// TIA Portal project "StepTimeAnalysis" (V16) (continued)
REGION Network 25: Archive values Step 9
   "DB_HMI".ARG1_Seq1_S9 := "IDB_Arg_Seq_1_DB".Step9.X;
END_REGION

REGION Network 26: Archive values Step 10
   "DB_HMI".ARG1_Seq1_S10 := "IDB_Arg_Seq_1_DB".Step10.X;
END_REGION

REGION Network 27: Archive values Step 11
   "DB_HMI".ARG1_Seq1_S11 := "IDB_Arg_Seq_1_DB".Step11.X;
END_REGION

REGION Network 28: Archive values Step 12
   "DB_HMI".ARG1_Seq1_S12 := "IDB_Arg_Seq_1_DB".Step12.X;
END_REGION

REGION Network 29: Archive values Step 13
   "DB_HMI".ARG1_Seq1_S13 := "IDB_Arg_Seq_1_DB".Step13.X;
END_REGION

REGION Network 30: Archive values Step 14
   "DB_HMI".ARG1_Seq1_S14 := "IDB_Arg_Seq_1_DB".Step14.X;
END_REGION

REGION Network 31: Archive values Step 15
   "DB_HMI".ARG1_Seq1_S15 := "IDB_Arg_Seq_1_DB".Step15.X;
END_REGION

REGION Network 32: Archive values Step 16
   "DB_HMI".ARG1_Seq1_S16 := "IDB_Arg_Seq_1_DB".Step16.X;
END_REGION

REGION Network 33: Archive values Step 17
   "DB_HMI".ARG1_Seq1_S17 := "IDB_Arg_Seq_1_DB".Step17.X;
END_REGION

REGION Network 34: Archive values Step 18
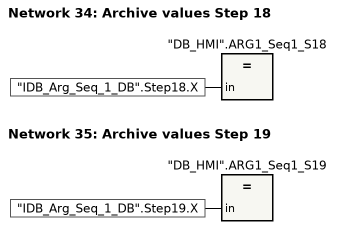
   "DB_HMI".ARG1_Seq1_S18 := "IDB_Arg_Seq_1_DB".Step18.X;
END_REGION

REGION Network 35: Archive values Step 19
   "DB_HMI".ARG1_Seq1_S19 := "IDB_Arg_Seq_1_DB".Step19.X;
END_REGION

REGION Network 36 (SCL): Set Busy
   IF
       "IDB_Arg_Seq_1_DB".Step2.X OR
       "IDB_Arg_Seq_1_DB".Step3.X OR
       "IDB_Arg_Seq_1_DB".Step4.X OR
       "IDB_Arg_Seq_1_DB".Step5.X OR
       "IDB_Arg_Seq_1_DB".Step6.X OR
       "IDB_Arg_Seq_1_DB".Step7.X OR
       "IDB_Arg_Seq_1_DB".Step8.X OR
       "IDB_Arg_Seq_1_DB".Step9.X OR
       "IDB_Arg_Seq_1_DB".Step10.X OR
       "IDB_Arg_Seq_1_DB".Step11.X OR
       "IDB_Arg_Seq_1_DB".Step12.X OR
       "IDB_Arg_Seq_1_DB".Step13.X OR
       "IDB_Arg_Seq_1_DB".Step14.X OR
       "IDB_Arg_Seq_1_DB".Step15.X OR
       "IDB_Arg_Seq_1_DB".Step16.X OR
       "IDB_Arg_Seq_1_DB".Step17.X OR
       "IDB_Arg_Seq_1_DB".Step18.X OR
       "IDB_Arg_Seq_1_DB".Step19.X THEN
       "DB_HMI".ARG1_Seq1_Status_Busy := TRUE;
   ELSIF "IDB_Arg_Seq_1_DB"."Step1: Init (Idle)".X THEN
       "DB_HMI".ARG1_Seq1_Status_Busy := FALSE;
   END_IF;
END_REGION

REGION Network 37 (SCL): When Stepper Sequence runs completely
   IF "IDB_Arg_Seq_1_DB".Trans10.TS = TRUE OR "IDB_Arg_Seq_1_DB".Trans21.TS = TRUE THEN
       "DB_Process_Var".Branch_Complete := TRUE;
       "DB_Process_Var".Car_Type_Ready := "DB_Process_Var".Car_Type_inProduction;
       "DB_Process_Var".Car_Type_inProduction := 0;
       "DB_Process_Var".Car_Type_inProduction_Text := '';
       "DB_Process_Var".Car_ReadyToShift := TRUE;
       "DB_HMI".ARG1_Seq1_inProduction := 0;
   END_IF;
   IF "IDB_Arg_Seq_1_DB".Trans1.TS = TRUE OR "IDB_Arg_Seq_1_DB".Trans11.TS = TRUE THEN
       "DB_Process_Var".Branch_Complete := FALSE;
       "DB_Process_Var".ReadyNewCar := 0;
   END_IF;
END_REGION

REGION Network 38 (SCL): Write Data in the Sending Box
   //IF "DB_Process_Var".Branch_Complete = TRUE AND "DB_PLC1_Receiving".ReceivingBox.Station_Idle = TRUE THEN
   IF "IDB_Arg_Seq_1_DB".Trans10.TS = TRUE OR "IDB_Arg_Seq_1_DB".Trans21.TS = TRUE THEN
       "DB_PLC1_Sending".SendBoxForward.Planned_PT_Red := "DB_HMI".ARG1_Seq1_Calculated_PT_Red;
       "DB_PLC1_Sending".SendBoxForward.Planned_PT_Green := "DB_HMI".ARG1_Seq1_Calculated_PT_Green;
       "DB_PLC1_Sending".SendBoxForward.Planned_PT_Blue := "DB_HMI".ARG1_Seq1_Calculated_PT_Blue;

       "DB_PLC1_Sending".SendBoxForward.Measuered_PT_Red := "DB_HMI".ARG1_Seq1_Messured_PT_Red;
       "DB_PLC1_Sending".SendBoxForward.Measuered_PT_Green := "DB_HMI".ARG1_Seq1_Messured_PT_Green;
       "DB_PLC1_Sending".SendBoxForward.Measuered_PT_Blue := "DB_HMI".ARG1_Seq1_Messured_PT_Blue;

       "DB_PLC1_Sending".SendBoxForward.Type := "DB_Process_Var".Car_Type_Ready;

       "DB_PLC1_Receiving".ReceivingBoxForward.Type := 0;
   END_IF;
END_REGION

REGION Network 39 (SCL)
   //IF "DB_Process_Var".Branch_Complete = TRUE AND "DB_PLC1_Receiving".ReceivingBox.Station_Idle = TRUE THEN
    //   "DB_Process_Var".ready_new_car := TRUE;
   //END_IF;
END_REGION

REGION Network 40 (SCL): When car is shifted
   IF "DB_Process_Var".Data_Put_Done = TRUE THEN
       "DB_Process_Var".Car_Type_Ready := 0;
       "DB_PLC1_Sending".SendBoxForward.Type := 0;
       "DB_Process_Var".Car_ReadyToShift := FALSE;
       "DB_Process_Var".ReadyNewCar := 1;

       //"DB_PLC1_Receiving".ReceivingBoxForward.Type := 0;
   END_IF;
END_REGION
END_FUNCTION

FUNCTION "FC_Com" : Void   // FC2, FBD
{ S7_Optimized_Access := 'TRUE' }
VERSION : 0.1
BEGIN

REGION Network 1: Communication PLC1 -> PLC2
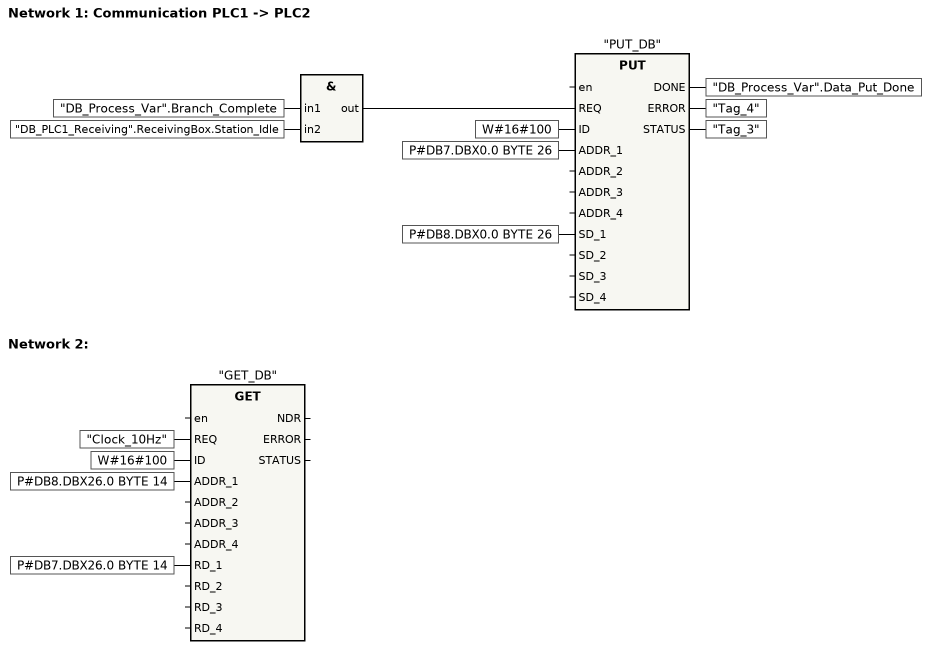
   "PUT_DB"(REQ := "DB_Process_Var".Branch_Complete AND "DB_PLC1_Receiving".ReceivingBox.Station_Idle,   // PUT
            ID := W#16#100,
            ADDR_1 := P#DB7.DBX0.0 BYTE 26,
            SD_1 := P#DB8.DBX0.0 BYTE 26,
            DONE => "DB_Process_Var".Data_Put_Done,
            ERROR => "Tag_4",
            STATUS => "Tag_3");
END_REGION

REGION Network 2
   "GET_DB"(REQ := "Clock_10Hz", ID := W#16#100, ADDR_1 := P#DB8.DBX26.0 BYTE 14, RD_1 := P#DB7.DBX26.0 BYTE 14);   // GET
END_REGION
END_FUNCTION

FUNCTION "FC_PT_Calc" : Void   // FC3, SCL
{ S7_Optimized_Access := 'TRUE' }
VERSION : 0.1
   VAR_TEMP
      i : Int;
   END_VAR
   VAR CONSTANT
      sequenceNO : Int := 9;
      Null : Time := T#0MS;
   END_VAR
BEGIN
   "DB_HMI".ARG1_Seq1_Calculated_PT_Red := #Null;
   "DB_HMI".ARG1_Seq1_Calculated_PT_Green := #Null;
   "DB_HMI".ARG1_Seq1_Calculated_PT_Blue := #Null;

   "DB_HMI".ARG1_Seq1_Messured_PT_Red := #Null;
   "DB_HMI".ARG1_Seq1_Messured_PT_Green := #Null;
   "DB_HMI".ARG1_Seq1_Messured_PT_Blue := #Null;

   FOR #i := 2 TO #sequenceNO + 1 DO
       //Calculated Production Time
       "DB_HMI".ARG1_Seq1_Calculated_PT_Red := "DB_HMI".ARG1_Seq1_Calculated_PT_Red + "DB_Profile".time_Red[#i];
       "DB_HMI".ARG1_Seq1_Calculated_PT_Green := "DB_HMI".ARG1_Seq1_Calculated_PT_Green + "DB_Profile".time_Green[#i];
       "DB_HMI".ARG1_Seq1_Calculated_PT_Blue := "DB_HMI".ARG1_Seq1_Calculated_PT_Blue + "DB_Profile".time_Blue[#i];
       //Messured Production Time
       IF "DB_Process_Var".Car_Type_inProduction = 3 THEN
           "DB_HMI".ARG1_Seq1_Messured_PT_Red := "DB_HMI".ARG1_Seq1_Messured_PT_Red + "DB_Process_Var".Step_Times[#i];
       ELSIF "DB_Process_Var".Car_Type_inProduction = 4 THEN
           "DB_HMI".ARG1_Seq1_Messured_PT_Green := "DB_HMI".ARG1_Seq1_Messured_PT_Green + "DB_Process_Var".Step_Times[#i];
       ELSIF "DB_Process_Var".Car_Type_inProduction = 6 THEN
           "DB_HMI".ARG1_Seq1_Messured_PT_Blue := "DB_HMI".ARG1_Seq1_Messured_PT_Blue + "DB_Process_Var".Step_Times[#i];
       END_IF;
   END_FOR;

   //Add Time of previous Stations
   "DB_HMI".ARG1_Seq1_Calculated_PT_Red := "DB_HMI".ARG1_Seq1_Calculated_PT_Red + "DB_PLC1_Receiving".ReceivingBoxForward.Planned_PT_Red;
   "DB_HMI".ARG1_Seq1_Calculated_PT_Green := "DB_HMI".ARG1_Seq1_Calculated_PT_Green + "DB_PLC1_Receiving".ReceivingBoxForward.Planned_PT_Green;
   "DB_HMI".ARG1_Seq1_Calculated_PT_Blue := "DB_HMI".ARG1_Seq1_Calculated_PT_Blue + "DB_PLC1_Receiving".ReceivingBoxForward.Planned_PT_Blue;

   "DB_HMI".ARG1_Seq1_Messured_PT_Red := "DB_HMI".ARG1_Seq1_Messured_PT_Red + "DB_PLC1_Receiving".ReceivingBoxForward.Measuered_PT_Red;
   "DB_HMI".ARG1_Seq1_Messured_PT_Green := "DB_HMI".ARG1_Seq1_Messured_PT_Green + "DB_PLC1_Receiving".ReceivingBoxForward.Measuered_PT_Green;
   "DB_HMI".ARG1_Seq1_Messured_PT_Blue := "DB_HMI".ARG1_Seq1_Messured_PT_Blue + "DB_PLC1_Receiving".ReceivingBoxForward.Measuered_PT_Blue;
END_FUNCTION

FUNCTION "FC_Global_Status" : Void   // FC4, SCL
{ S7_Optimized_Access := 'TRUE' }
VERSION : 0.1
   VAR_TEMP
      global_auto : Bool;
      global_man : Bool;
      test2 : Bool;
      test : Bool;
      i : Int;
   END_VAR
BEGIN
   IF "DB_Process_Var".Auto_Mode = TRUE THEN
       "DB_PLC1_Sending".SendBox.Mode_PLC1 := 1;
   ELSIF "DB_Process_Var".Man_Mode = TRUE THEN
       "DB_PLC1_Sending".SendBox.Mode_PLC1 := 2;
   ELSE
       "DB_PLC1_Sending".SendBox.Mode_PLC1 := 0;
   END_IF;

   IF "DB_Process_Var".Station_Nr = 1 THEN
       IF "DB_PLC1_Sending".SendBox.Mode_PLC1 = 1 AND "DB_PLC1_Receiving".ReceivingBox.Mode_PLC2 = 1 AND "DB_PLC1_Receiving".ReceivingBox.Mode_PLC3 = 1 AND "DB_PLC1_Receiving".ReceivingBox.Mode_PLC4 = 1 AND "DB_PLC1_Receiving".ReceivingBox.Mode_PLC5 = 1 THEN
           "DB_HMI".Global_Status_Auto := TRUE;
           "DB_HMI".Global_Status_Man := FALSE;
       ELSIF "DB_PLC1_Sending".SendBox.Mode_PLC1 = 0 AND "DB_PLC1_Receiving".ReceivingBox.Mode_PLC2 = 0 AND "DB_PLC1_Receiving".ReceivingBox.Mode_PLC3 = 0 AND "DB_PLC1_Receiving".ReceivingBox.Mode_PLC4 = 0 AND "DB_PLC1_Receiving".ReceivingBox.Mode_PLC5 = 0 THEN
           "DB_HMI".Global_Status_Auto := FALSE;
           "DB_HMI".Global_Status_Man := FALSE;
       ELSE
           "DB_HMI".Global_Status_Man := TRUE;
           "DB_HMI".Global_Status_Auto := FALSE;
       END_IF;
   END_IF;


   //Global Selection
   "DB_PLC1_Receiving".ReceivingBoxForward.Type := "DB_HMI".Global_selection;
END_FUNCTION

ORGANIZATION_BLOCK "Main"   // OB1, LAD, ProgramCycle
TITLE = "Main Program Sweep (Cycle)"
{ S7_Optimized_Access := 'TRUE' }
VERSION : 0.1
   VAR_INPUT
      Initial_Call : Bool;   // Initial call of this OB
      Remanence : Bool;   // =True, if remanent data are available
   END_VAR
   VAR_TEMP
      test : Bool;
   END_VAR
BEGIN

REGION Network 1: Call ARG_1
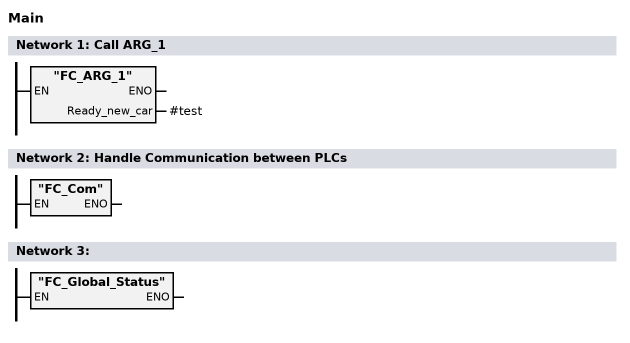
   RUNG wire#powerrail
      "FC_ARG_1"(Ready_new_car => #test)
   END_RUNG
   // the same network as SCL:
   "FC_ARG_1"(Ready_new_car => #test);
END_REGION

REGION Network 2: Handle Communication between PLCs
   RUNG wire#powerrail
      "FC_Com"()
   END_RUNG
   // the same network as SCL:
   "FC_Com"();
END_REGION

REGION Network 3
   RUNG wire#powerrail
      "FC_Global_Status"()
   END_RUNG
   // the same network as SCL:
   "FC_Global_Status"();
END_REGION
END_ORGANIZATION_BLOCK

// folder: LGF/4 Math operations

FUNCTION "LGF_RandomRange_Dint" : DInt   // FC10013, SCL
TITLE = LGF_RandomRange_DInt
{ S7_Optimized_Access := 'TRUE' }
AUTHOR : Siemens_Digital_Industries
FAMILY : LGF
NAME : LGF_RandomRange_DInt
// This function generates random numbers in defined limits (Datatype DInt)
   VAR_INPUT
      minValue : DInt;   // minimal Value random can reach / Minimum value of the range of the random number
      maxValue : DInt;   // maximal Value random can reach / Maximum value of the range of the random number
   END_VAR
   VAR_OUTPUT
      error : Bool;   // Error if true
      status : Word;   // Status of the function
      subfunctionStatus : Word;   // Status or return value of called FB's, FCs and system blocks
   END_VAR
   VAR_TEMP
      tempTime : DTL;   // System time
      tempNanoSecondInDWord : DWord;   // UDINT converted to DWORD for access to individual bytes
      tempTimeStatus : Word;   // Status of the instruction RD_SYS_T
      tempRandomValue : DWord;   // Random-start-value
      tempNormReal : Real;   // Normalized value
   END_VAR
   // Ret_Val : Returns random DInt number in a predefined range
   VAR CONSTANT
      ZERO : DInt := 0;   // Zero value in case of error
      MAX_UDINT : UDInt := 4294967295 ;   // Maximum UDINT value
      SUB_STATUS_NO_ERROR : Word := 16#0000;   // Status: sub function call ends without error
      STATUS_FINISHED_NO_ERROR : Word := 16#0000;   // Status: Execution finished without errors
      ERR_MAX_LESS_MIN : Word := 16#8200;   // Error: The maximum limit number is smaller than the minimum limit number
      ERR_RD_SYS_T : Word := 16#8600;   // Error: System function Read system time returned an error
   END_VAR
BEGIN
   REGION Block info header
     //=============================================================================
     // SIEMENS AG / (c)Copyright 2017
     //-----------------------------------------------------------------------------
     // Title:            LGF_RandomRange_DInt
     // Comment/Function: This function generates random numbers in defined limits (Datatype DInt)
     // Library/Family:   LGF(Library General Functions)
     // Author:           Siemens Digital Industry Support
     // Tested with:      S7-PLCSIM Advanced V2.0 SP1
     // Engineering:      TIA Portal V15 Update 2
     // Restrictions:     ENO disabled - error handling done by error and status
     // Requirements:     PLC (S7-1200 / S7-1500)
     //-------------------------------------------------------------------------------
     // Change log table:
     // Version  | Date       | Expert in charge       | Changes applied
     //----------|------------|------------------------|------------------------------
     // 01.00.00 19.08.2015  Siemens Industry Online Support
     //                      First released version
     // 01.00.01 02.01.2017  Siemens Industry Online Support
     //                      Upgrade: TIA Portal V14 Update 1
     // 01.00.02 17.08.2018  Siemens Industry Online Support
     //                      Upgrade: TIA V15 Update 2
     // 01.00.03 23.11.2018  Siemens Industry Online Support
     //                      Upgrade: TIA V15.1
     // 01.01.00 09.10.2019  Siemens Industry Presales Support
     //                      Renamed from "LGF_RandomInt" to "LGF_RandomRange_DInt"
     //                      change random datatype from int to dint
     //                      Regions, commens and costants are added
     // 03.00.00 23.04.2020  Siemens Industry Support
     //                      Set version to V3.0.0, harmonize the version of the whole library
     //=============================================================================
   END_REGION

   REGION Validation
     // Check if the maximal Value is less than the minimal value
     IF (#minValue > #maxValue) THEN
       #error := true;
       #status := #ERR_MAX_LESS_MIN;
       #subfunctionStatus := #SUB_STATUS_NO_ERROR;
       #LGF_RandomRange_Dint := #ZERO;
       RETURN;
     END_IF;

     // Read system time
     #tempTimeStatus := INT_TO_WORD(RD_SYS_T(#tempTime));

     // Check return variable for error
     IF (#tempTimeStatus <> #SUB_STATUS_NO_ERROR) THEN
       #error := true;
       #status := #ERR_RD_SYS_T;
       #subfunctionStatus := #tempTimeStatus;
       #LGF_RandomRange_Dint := #ZERO;
       RETURN;
     END_IF;
   END_REGION

   REGION Calculating random number
     // Converting to double word so individual bytes can be addressed
     #tempNanoSecondInDWord := UDINT_TO_DWORD(#tempTime.NANOSECOND);

     // Callculate a random-start-value depending on the time
     #tempRandomValue.%B3 := #tempNanoSecondInDWord.%B0;
     #tempRandomValue.%B2 := #tempNanoSecondInDWord.%B1;
     #tempRandomValue.%B1 := #tempNanoSecondInDWord.%B2;
     #tempRandomValue.%B0 := #tempNanoSecondInDWord.%B3;

     // Norm the calculated random number: 0.0 <= #tempNormReal <= 1.0
     #tempNormReal := UDINT_TO_REAL(DWORD_TO_UDINT(#tempRandomValue)) / UDINT_TO_REAL(#MAX_UDINT);

     // Scale the tempNormReal to be in the range of maxValue and minValue
     #LGF_RandomRange_Dint := REAL_TO_DINT((#tempNormReal * DINT_TO_REAL(#maxValue - #minValue) + DINT_TO_REAL(#minValue)));

     #error := false;
     #status := #STATUS_FINISHED_NO_ERROR;
     #subfunctionStatus := #SUB_STATUS_NO_ERROR;
     // ENO mechanism is not used
     ENO := TRUE;
   END_REGION
END_FUNCTION

FUNCTION "LGF_Random_DInt" : DInt   // FC10084, SCL
TITLE = LGF_Random_DInt
{ S7_Optimized_Access := 'TRUE' }
AUTHOR : Siemens_Digital_Industries
FAMILY : LGF
NAME : LGF_Random_DInt
// Generates a random number in the DInt Range
   VAR_OUTPUT
      error : Bool;   // Error if true
      status : Word;   // Status of the function
      subfunctionStatus : Word;   // Status or return value of called FB's, FCs and system blocks
   END_VAR
   VAR_TEMP
      tempTime : DTL;   // System time
      tempNanoSecondInDWord : DWord;   // UDINT converted to DWORD for access to individual bytes
      tempTimeStatus : Word;   // Status of the instruction RD_SYS_T
      tempRandomValue : DWord;   // Random-start-value
   END_VAR
   // Ret_Val : Random number in the Dint range
   VAR CONSTANT
      ZERO : DInt;   // Zero value in case of error
      SUB_STATUS_NO_ERROR : Word := 16#0000;   // Status: sub function call ends without error
      STATUS_FINISHED_NO_ERROR : Word := 16#0000;   // Status: Execution finished without errors
      ERR_RD_SYS_T : Word := 16#8600;   // Error: System function Read system time returned an error
   END_VAR
BEGIN
   REGION Block info header
     //=============================================================================
     // SIEMENS AG / (c)Copyright 2017
     //-----------------------------------------------------------------------------
     // Title:            LGF_Random_DInt
     // Comment/Function: Generates a random number in the DInt Range
     // Library/Family:   LGF(Library General Functions)
     // Author:           Siemens Digital Industry Support
     // Tested with:      S7-PLCSIM Advanced V2.0 SP1
     // Engineering:      TIA Portal V15 Update 2
     // Restrictions:     ENO disabled - error handling done by error and status
     // Requirements:     PLC (S7-1200 / S7-1500)
     //-------------------------------------------------------------------------------
     // Change log table:
     // Version  | Date       | Expert in charge       | Changes applied
     //----------|------------|------------------------|------------------------------
     // 01.00.00 13.11.2019  Siemens Industry Presales Support
     //                      First release
     //                      copied from "LGF_Random_Real"
     // 03.00.00 23.04.2020  Siemens Industry Support
     //                      Set version to V3.0.0, harmonize the version of the whole library
     //=============================================================================
   END_REGION

   REGION Validation
     // Read system time
     #tempTimeStatus := INT_TO_WORD(RD_SYS_T(#tempTime));

     // Check return variable for error
     IF (#tempTimeStatus <> #SUB_STATUS_NO_ERROR) THEN
       #error := true;
       #status := #ERR_RD_SYS_T;
       #subfunctionStatus := #tempTimeStatus;
       #LGF_Random_DInt := #ZERO;
       RETURN;
     END_IF;
   END_REGION

   REGION Calculating random number
     // Converting to double word so individual bytes can be addressed
     #tempNanoSecondInDWord := UDINT_TO_DWORD(#tempTime.NANOSECOND);

     // Calculate a random-start-value depending on the time
     #tempRandomValue.%B3 := #tempNanoSecondInDWord.%B0;
     #tempRandomValue.%B2 := #tempNanoSecondInDWord.%B1;
     #tempRandomValue.%B1 := #tempNanoSecondInDWord.%B2;
     #tempRandomValue.%B0 := #tempNanoSecondInDWord.%B3;

     #LGF_Random_DInt := DWORD_TO_DINT(#tempRandomValue);

     #error := false;
     #status := #STATUS_FINISHED_NO_ERROR;
     #subfunctionStatus := #SUB_STATUS_NO_ERROR;
     // ENO mechanism is not used
     ENO := TRUE;
   END_REGION
END_FUNCTION

// ===== PLC "PLC_2"  CPU 1518F-4 PN/DP =====

VAR_GLOBAL   // PLC tag table "Default tag table"
   "Clock_Byte" AT %MB0 : Byte;
   "Clock_10Hz" AT %M0.0 : Bool;
   "Clock_5Hz" AT %M0.1 : Bool;
   "Clock_2.5Hz" AT %M0.2 : Bool;
   "Clock_2Hz" AT %M0.3 : Bool;
   "Clock_1.25Hz" AT %M0.4 : Bool;
   "Clock_1Hz" AT %M0.5 : Bool;
   "Clock_0.625Hz" AT %M0.6 : Bool;
   "Clock_0.5Hz" AT %M0.7 : Bool;
   "Tag_1" AT %M10.1 : Bool;
   "Tag_2" AT %M10.2 : Bool;
   "Tag_3" AT %MW14 : Word;
END_VAR

TYPE "PLC_SF"
   STRUCT
      "Type" : Int;
      Planned_PT_Red : Time;
      Planned_PT_Green : Time;
      Planned_PT_Blue : Time;
      Measuered_PT_Red : Time;
      Measuered_PT_Green : Time;
      Measuered_PT_Blue : Time;
   END_STRUCT;
END_TYPE

TYPE "PLC_SR"
   STRUCT
      "Type" : Int;
      Station_Idle : Bool;
      Mode_PLC1 : Int;
      Mode_PLC2 : Int;
      Mode_PLC3 : Int;
      Mode_PLC4 : Int;
      Mode_PLC5 : Int;
   END_STRUCT;
END_TYPE

DATA_BLOCK "IDB_Arg_Seq_1_DB"   // DB2
{ S7_Optimized_Access := 'TRUE' }
VERSION : 0.1
// stored: InstanceOfName FB_Arg_Seq_1
"FB_Arg_Seq_1"
BEGIN
END_DATA_BLOCK

DATA_BLOCK "DB_HMI"   // DB3
{ S7_Optimized_Access := 'TRUE' }
VERSION : 0.1
   VAR
      ARG1_Seq1_S1 : Bool;
      ARG1_Seq1_T1 : Bool;
      ARG1_Seq1_S2 : Bool;
      ARG1_Seq1_T2 : Bool;
      ARG1_Seq1_S3 : Bool;
      ARG1_Seq1_T3 : Bool;
      ARG1_Seq1_S4 : Bool;
      ARG1_Seq1_T4 : Bool;
      ARG1_Seq1_S5 : Bool;
      ARG1_Seq1_T5 : Bool;
      ARG1_Seq1_S6 : Bool;
      ARG1_Seq1_T6 : Bool;
      ARG1_Seq1_S7 : Bool;
      ARG1_Seq1_T7 : Bool;
      ARG1_Seq1_S8 : Bool;
      ARG1_Seq1_T8 : Bool;
      ARG1_Seq1_S9 : Bool;
      ARG1_Seq1_T9 : Bool;
      ARG1_Seq1_S10 : Bool;
      ARG1_Seq1_T10 : Bool;
      ARG1_Seq1_S11 : Bool;
      ARG1_Seq1_T11 : Bool;
      ARG1_Seq1_S12 : Bool;
      ARG1_Seq1_T12 : Bool;
      ARG1_Seq1_S13 : Bool;
      ARG1_Seq1_T13 : Bool;
      ARG1_Seq1_S14 : Bool;
      ARG1_Seq1_T14 : Bool;
      ARG1_Seq1_S15 : Bool;
      ARG1_Seq1_T15 : Bool;
      ARG1_Seq1_S16 : Bool;
      ARG1_Seq1_T16 : Bool;
      ARG1_Seq1_S17 : Bool;
      ARG1_Seq1_T17 : Bool;
      ARG1_Seq1_S18 : Bool;
      ARG1_Seq1_T18 : Bool;
      ARG1_Seq1_S19 : Bool;
      ARG1_Seq1_T19 : Bool;
      inputTimes : Array[2..10] of DInt;
      dropdown_selection : Int := 3;
      ARG1_Seq1_Status_Idle : Bool;   // Stepper Sequence is in Idle (Step 1)
      ARG1_Seq1_Status_Busy : Bool;   // Stepper Stequence is Busy (Step2 - Step 19)
      ARG1_Seq1_Status_Man : Bool;   // Status Stepper Sequence is in Manuel Mode
      ARG1_Seq1_Status_Auto : Bool;   // Status Stepper Sequence is in Auto Mode
      ARG1_Seq1_Cmd_Man : Bool;   // Command Manuel Mode for Stepper Sequence
      ARG1_Seq1_Cmd_Auto : Bool;   // Command Auto Mode for Stepper Sequence
      ARG1_Seq1_Cmd_Stop : Bool;   // Command Stop for Stepper Sequence
      ARG1_Seq1_Cmd_Start : Bool;   // Command Start for Stepper Sequence
      ARG1_Seq1_Cmd_DelayReset : Bool;
      Global_Cmd_Auto : Bool;
      Global_Cmd_Man : Bool;
      Global_Cmd_Start : Bool;
      Global_Cmd_Stop : Bool;
      Global_Status_Man : Bool;
      Global_Status_Auto : Bool;
      Global_selection : Int;
      ARG1_Seq1_inProduction : Int;
      ARG1_Seq1_Calculated_PT_Red : Time;
      ARG1_Seq1_Calculated_PT_Green : Time;
      ARG1_Seq1_Calculated_PT_Blue : Time;
      ARG1_Seq1_Messured_PT_Red : Time;
      ARG1_Seq1_Messured_PT_Green : Time;
      ARG1_Seq1_Messured_PT_Blue : Time;
      ARG1_Seq1_DelaySelect_Red : Array[2..10] of Bool;
      ARG1_Seq1_DelaySelect_Green : Array[2..10] of Bool;
      ARG1_Seq1_DelaySelect_Blue : Array[2..10] of Bool;
   END_VAR
BEGIN
END_DATA_BLOCK

DATA_BLOCK "DB_Sim"   // DB4
{ S7_Optimized_Access := 'TRUE' }
VERSION : 0.1
   VAR
      Delta_T_Red : Array[2..10] of Time;
      Delta_T_Green : Array[2..10] of Time;
      Delta_T_Blue : Array[2..10] of Time;
   END_VAR
BEGIN
   Delta_T_Red[2] := T#100ms;
   Delta_T_Red[3] := T#100ms;
   Delta_T_Red[4] := T#100ms;
   Delta_T_Red[5] := T#100ms;
   Delta_T_Red[6] := T#100ms;
   Delta_T_Red[7] := T#100ms;
   Delta_T_Red[8] := T#100ms;
   Delta_T_Red[9] := T#100ms;
   Delta_T_Red[10] := T#100ms;
END_DATA_BLOCK

DATA_BLOCK "DB_Profile"   // DB5
{ S7_Optimized_Access := 'TRUE' }
VERSION : 0.1
   VAR
      "time" : Array[2..10] of Time;
      time_Red : Array[2..10] of Time;
      time_Green : Array[2..10] of Time;
      time_Blue : Array[2..10] of Time;
   END_VAR
BEGIN
   time_Red[2] := t#3s;
   "time"[2] := t#3s;
   "time"[3] := t#3s;
   "time"[4] := t#3s;
   "time"[5] := t#3s;
   "time"[6] := t#3s;
   "time"[7] := t#3s;
   "time"[8] := t#3s;
   "time"[9] := t#3s;
   "time"[10] := t#3s;
   time_Red[3] := t#6s;
   time_Red[4] := t#5s;
   time_Red[5] := t#9s;
   time_Red[6] := t#4s;
   time_Red[7] := t#6s;
   time_Red[8] := t#8s;
   time_Red[9] := t#7s;
   time_Red[10] := t#4s;
   time_Green[2] := t#7s;
   time_Green[3] := t#4s;
   time_Green[4] := t#8s;
   time_Green[5] := t#4s;
   time_Green[6] := t#3s;
   time_Green[7] := t#9s;
   time_Green[8] := t#5s;
   time_Green[9] := t#6s;
   time_Green[10] := t#8s;
   time_Blue[2] := t#4s;
   time_Blue[3] := t#6s;
   time_Blue[4] := t#9s;
   time_Blue[5] := t#3s;
   time_Blue[6] := t#7s;
   time_Blue[7] := t#6s;
   time_Blue[8] := t#5s;
   time_Blue[9] := t#9s;
   time_Blue[10] := t#6s;
END_DATA_BLOCK

DATA_BLOCK "DB_Process_Var"   // DB6
{ S7_Optimized_Access := 'TRUE' }
VERSION : 0.1
   VAR
      Man_Mode : Bool := true;
      Auto_Mode : Bool;
      Start : Bool;
      Branch_Complete : Bool;
      Step_Times : Array[2..10] of Time;
      Car_Type_Selected : Int;
      Car_Type_inProduction : Int;
      Car_Type_Ready : Int;
      Car_ReadyToShift : Bool;
      Data_Put_Done : Bool;
      Car_Type_inProduction_Text : String;
      Station_Nr : Int := 2;
      ReadyNewCar : Bool := true;
      Global_Start : Bool;
      Global_Stop : Bool;
   END_VAR
BEGIN
END_DATA_BLOCK

DATA_BLOCK "DB_PLC2_Receiving"   // DB7
{ S7_Optimized_Access := 'FALSE' }
VERSION : 0.1
   VAR
      ReceivingBoxForward : "PLC_SF";
      ReceivingBox : "PLC_SR";
   END_VAR
BEGIN
END_DATA_BLOCK

DATA_BLOCK "DB_PLC2_Sending"   // DB8
{ S7_Optimized_Access := 'FALSE' }
VERSION : 0.1
   VAR
      SendBoxForward : "PLC_SF";
      SendBox : "PLC_SR";
   END_VAR
BEGIN
END_DATA_BLOCK

FUNCTION_BLOCK "FB_Arg_Seq_1"   // FB2, GRAPH_PLUS
{ S7_Optimized_Access := 'TRUE' }
VERSION : 0.1
   VAR_INPUT
      OFF_SQ : Bool := false;   // Turn sequence off
      INIT_SQ : Bool := false;   // Set sequence to initial state
      ACK_EF : Bool := false;   // Acknowledge all errors and faults
      S_PREV : Bool := false;   // Output previous step in parameter S_NO
      S_NEXT : Bool := false;   // Indicate next step in parameter S_NO
      SW_AUTO : Bool := false;   // Automatic mode
      SW_TAP : Bool := false;   // Semiautomatic/switch with transition
      SW_TOP : Bool := false;   // Semiautomatic/ignore transition
      SW_MAN : Bool := false;   // Manual mode
      S_SEL : Int := 0;   // Select step to be output to S_NO
      S_ON : Bool := false;   // Activate step indicated in S_NO
      S_OFF : Bool := false;   // Deactivate step indicated S_NO
      T_PUSH : Bool := false;   // Enable transition to switch in semi automatic mode
      Start : Bool;
      stepTimes : Array[2..10] of Time;
      Model_Numb : Int := 3;
   END_VAR
   VAR_OUTPUT
      S_NO : Int := 0;   // Step number
      S_MORE : Bool := false;   // More steps are available and can be shown in S_NO
      S_ACTIVE : Bool := false;   // Step indicated in S_NO is active
      ERR_FLT : Bool := false;   // Interlock or supervision group error
      AUTO_ON : Bool := false;   // Automatic mode is active
      TAP_ON : Bool := false;   // Semiautomatic mode/step with transition enabled
      TOP_ON : Bool := false;   // Semiautomatic mode/ignore transition enabled
      MAN_ON : Bool := false;   // Manual mode is active
   END_VAR
   VAR
      HMI_INFO : Array[0..8] of UInt;
      IF_PAR : G7_IfParPlus_V6;
      RT_DATA : G7_RTDataPlus_V6;   // Internal data area
      Trans1 : G7_TransitionPlus_V6;   // Transition structure
      Trans2 : G7_TransitionPlus_V6;   // Transition structure
      Trans3 : G7_TransitionPlus_V6;   // Transition structure
      Trans4 : G7_TransitionPlus_V6;   // Transition structure
      Trans5 : G7_TransitionPlus_V6;   // Transition structure
      Trans6 : G7_TransitionPlus_V6;   // Transition structure
      Trans7 : G7_TransitionPlus_V6;   // Transition structure
      Trans8 : G7_TransitionPlus_V6;   // Transition structure
      Trans9 : G7_TransitionPlus_V6;   // Transition structure
      Trans10 : G7_TransitionPlus_V6;   // Transition structure
      Trans11 : G7_TransitionPlus_V6;   // Transition structure
      Trans12 : G7_TransitionPlus_V6;   // Transition structure
      Trans13 : G7_TransitionPlus_V6;   // Transition structure
      Trans14 : G7_TransitionPlus_V6;   // Transition structure
      Trans15 : G7_TransitionPlus_V6;   // Transition structure
      Trans16 : G7_TransitionPlus_V6;   // Transition structure
      Trans17 : G7_TransitionPlus_V6;   // Transition structure
      Trans18 : G7_TransitionPlus_V6;   // Transition structure
      Trans19 : G7_TransitionPlus_V6;   // Transition structure
      Trans21 : G7_TransitionPlus_V6;   // Transition structure
      "Step1: Init (Idle)" : G7_StepPlus_V6;   // Step structure
      Step2 : G7_StepPlus_V6;   // Step structure
      Step3 : G7_StepPlus_V6;   // Step structure
      Step4 : G7_StepPlus_V6;   // Step structure
      Step5 : G7_StepPlus_V6;   // Step structure
      Step6 : G7_StepPlus_V6;   // Step structure
      Step7 : G7_StepPlus_V6;   // Step structure
      Step8 : G7_StepPlus_V6;   // Step structure
      Step9 : G7_StepPlus_V6;   // Step structure
      Step10 : G7_StepPlus_V6;   // Step structure
      Step11 : G7_StepPlus_V6;   // Step structure
      Step12 : G7_StepPlus_V6;   // Step structure
      Step13 : G7_StepPlus_V6;   // Step structure
      Step14 : G7_StepPlus_V6;   // Step structure
      Step15 : G7_StepPlus_V6;   // Step structure
      Step16 : G7_StepPlus_V6;   // Step structure
      Step17 : G7_StepPlus_V6;   // Step structure
      Step18 : G7_StepPlus_V6;   // Step structure
      Step19 : G7_StepPlus_V6;   // Step structure
      SINI : Array[0..1] of USInt;
      LSTT : Array[0..19] of USInt;
      ATAJ : Array[0..19] of USInt;
      ATAB : Array[0..19] of USInt;
      PSTT : Array[0..19] of USInt;
      NSTT : Array[0..19] of USInt;
      ASSJ : Array[0..18] of USInt;
      ASSB : Array[0..18] of USInt;
      PTTS : Array[0..18] of USInt;
      NTTS : Array[0..18] of USInt;
      SW_SQTS : Array[0..18] of USInt;
      SWITCH : Array[0..1] of USInt;
      TVX : Array[0..3] of USInt;
      TTX : Array[0..3] of USInt;
      TSX : Array[0..1] of USInt;
      S00X : Array[0..1] of USInt;
      SOFFX : Array[0..1] of USInt;
      SONX : Array[0..1] of USInt;
      SAX : Array[0..1] of USInt;
      SERRX : Array[0..19] of USInt;
      SMX : Array[0..19] of USInt;
      S0X : Array[0..19] of USInt;
      S1X : Array[0..19] of USInt;
      IL_ALARM_INST : Diag_Alarm;
      SUP_ALARM_INST : Diag_Alarm;
      STEP_TIME_ALARM_INST : Diag_Alarm;
      IEC_TIMER_INST : IEC_TIMER;
      TRANSACTION_FLAG : Bool := false;
   END_VAR
   // SINI[0] := 2;
   // LSTT[0] := 255;
   // LSTT[1] := 255;
   // LSTT[2] := 255;
   // ATAJ[1] := 1;
   // ATAJ[2] := 2;
   // ATAJ[3] := 3;
   // ATAB[1] := 1;
   // ATAB[2] := 2;
   // ATAB[3] := 3;
   // PSTT[1] := 1;
   // PSTT[2] := 2;
   // PSTT[3] := 3;
   // NSTT[0] := 1;
   // NSTT[1] := 2;
   // NSTT[2] := 3;
   // ASSJ[1] := 1;
   // ASSJ[2] := 2;
   // ASSJ[3] := 3;
   // ASSB[1] := 1;
   // ASSB[2] := 2;
   // ASSB[3] := 3;
   // PTTS[0] := 255;
   // PTTS[2] := 1;
   // PTTS[3] := 2;
   // NTTS[1] := 1;
   // NTTS[2] := 2;
   // NTTS[3] := 3;
   // TVX[0] := 16#1;
   // TTX[0] := 16#1;
   // TSX[0] := 16#1;
   // S00X[0] := 16#1;
   // SOFFX[0] := 16#1;
   // SONX[0] := 16#1;
   // SAX[0] := 16#1;
   // SERRX[0] := 16#1;
   // SMX[0] := 16#1;
   // S0X[0] := 16#1;
   // S1X[0] := 16#1;
   // LSTT[3] := 255;
   // LSTT[4] := 255;
   // LSTT[5] := 255;
   // LSTT[6] := 255;
   // LSTT[7] := 255;
   // LSTT[8] := 255;
   // ATAJ[4] := 4;
   // ATAJ[5] := 5;
   // ATAJ[6] := 6;
   // ATAJ[7] := 7;
   // ATAJ[8] := 8;
   // ATAJ[9] := 9;
   // ATAB[4] := 4;
   // ATAB[5] := 5;
   // ATAB[6] := 6;
   // ATAB[7] := 7;
   // ATAB[8] := 8;
   // ATAB[9] := 9;
   // PSTT[4] := 4;
   // PSTT[5] := 5;
   // PSTT[6] := 6;
   // PSTT[7] := 7;
   // PSTT[8] := 8;
   // PSTT[9] := 9;
   // NSTT[3] := 4;
   // NSTT[4] := 5;
   // NSTT[5] := 6;
   // NSTT[6] := 7;
   // NSTT[7] := 8;
   // NSTT[8] := 9;
   // ASSJ[4] := 4;
   // ASSJ[5] := 5;
   // ASSJ[6] := 6;
   // ASSJ[7] := 7;
   // ASSJ[8] := 8;
   // ASSJ[9] := 9;
   // ASSB[4] := 4;
   // ASSB[5] := 5;
   // ASSB[6] := 6;
   // ASSB[7] := 7;
   // ASSB[8] := 8;
   // ASSB[9] := 9;
   // PTTS[4] := 3;
   // PTTS[5] := 4;
   // PTTS[6] := 5;
   // PTTS[7] := 6;
   // PTTS[8] := 7;
   // PTTS[9] := 8;
   // NTTS[4] := 4;
   // NTTS[5] := 5;
   // NTTS[6] := 6;
   // NTTS[7] := 7;
   // NTTS[8] := 8;
   // NTTS[9] := 9;
   // LSTT[10] := 255;
   // LSTT[11] := 255;
   // LSTT[12] := 255;
   // LSTT[13] := 255;
   // LSTT[14] := 255;
   // LSTT[15] := 255;
   // LSTT[16] := 255;
   // LSTT[17] := 255;
   // LSTT[18] := 255;
   // ATAJ[10] := 10;
   // ATAJ[11] := 11;
   // ATAJ[12] := 12;
   // ATAJ[13] := 13;
   // ATAJ[14] := 14;
   // ATAJ[15] := 15;
   // ATAJ[16] := 16;
   // ATAJ[17] := 17;
   // ATAJ[18] := 18;
   // ATAJ[19] := 19;
   // ATAB[0] := 10;
   // ATAB[11] := 11;
   // ATAB[12] := 12;
   // ATAB[13] := 13;
   // ATAB[14] := 14;
   // ATAB[15] := 15;
   // ATAB[16] := 16;
   // ATAB[17] := 17;
   // ATAB[18] := 18;
   // ATAB[19] := 19;
   // PSTT[11] := 10;
   // PSTT[12] := 11;
   // PSTT[13] := 12;
   // PSTT[14] := 13;
   // PSTT[15] := 14;
   // PSTT[16] := 15;
   // PSTT[17] := 16;
   // PSTT[18] := 17;
   // PSTT[19] := 18;
   // NSTT[10] := 10;
   // NSTT[11] := 11;
   // NSTT[12] := 12;
   // NSTT[13] := 13;
   // NSTT[14] := 14;
   // NSTT[15] := 15;
   // NSTT[16] := 16;
   // NSTT[17] := 17;
   // NSTT[18] := 18;
   // ASSJ[10] := 10;
   // ASSJ[11] := 11;
   // ASSJ[12] := 12;
   // ASSJ[13] := 13;
   // ASSJ[14] := 14;
   // ASSJ[15] := 15;
   // ASSJ[16] := 16;
   // ASSJ[17] := 17;
   // ASSJ[18] := 18;
   // ASSB[10] := 10;
   // ASSB[11] := 11;
   // ASSB[12] := 12;
   // ASSB[13] := 13;
   // ASSB[14] := 14;
   // ASSB[15] := 15;
   // ASSB[16] := 16;
   // ASSB[17] := 17;
   // ASSB[18] := 18;
   // PTTS[10] := 10;
   // PTTS[11] := 11;
   // PTTS[12] := 12;
   // PTTS[13] := 13;
   // PTTS[14] := 14;
   // PTTS[15] := 15;
   // PTTS[16] := 16;
   // PTTS[17] := 17;
   // PTTS[18] := 18;
   // NTTS[10] := 11;
   // NTTS[11] := 12;
   // NTTS[12] := 13;
   // NTTS[13] := 14;
   // NTTS[14] := 15;
   // NTTS[15] := 16;
   // NTTS[16] := 17;
   // NTTS[17] := 18;
   // NTTS[18] := 19;
   // SW_SQTS[1] := 1;
   // SW_SQTS[2] := 1;
   // SW_SQTS[3] := 1;
   // SW_SQTS[4] := 1;
   // SW_SQTS[5] := 1;
   // SW_SQTS[6] := 1;
   // SW_SQTS[7] := 1;
   // SW_SQTS[8] := 1;
   // SW_SQTS[9] := 1;
   // SW_SQTS[10] := 2;
   // SW_SQTS[11] := 2;
   // SW_SQTS[12] := 2;
   // SW_SQTS[13] := 2;
   // SW_SQTS[14] := 2;
   // SW_SQTS[15] := 2;
   // SW_SQTS[16] := 2;
   // SW_SQTS[17] := 2;
   // SW_SQTS[18] := 2;
BEGIN